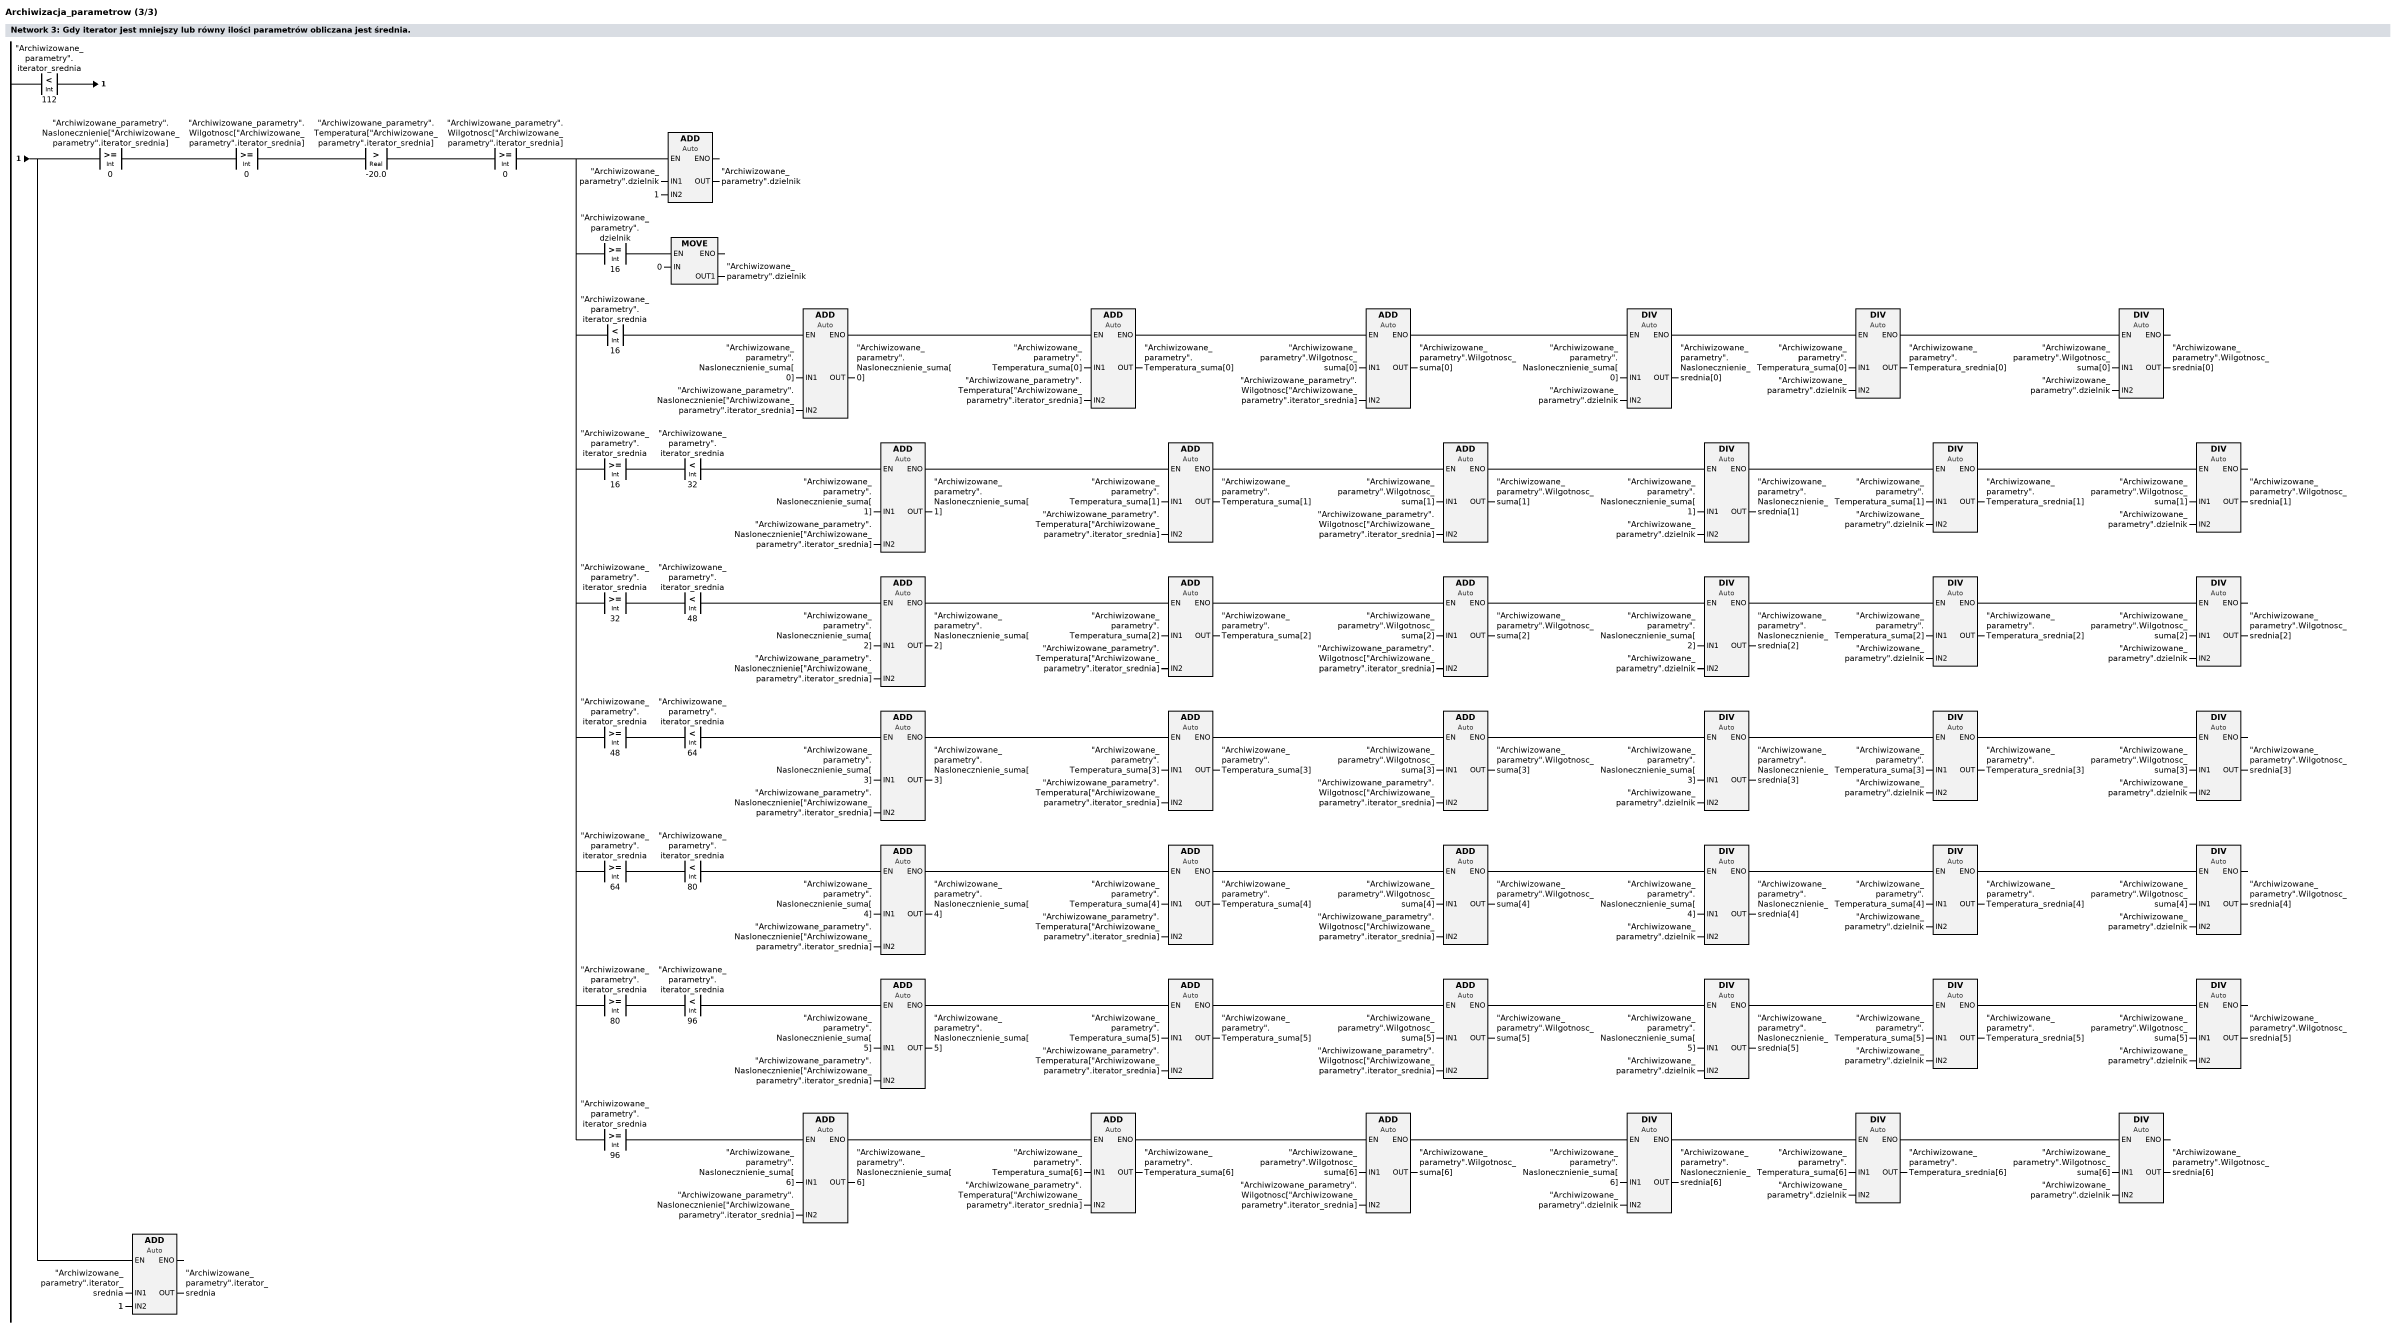
   RUNG wire#powerrail
      { S7_Templates := "SrcType := Int" } LT_Contact(in1 := "Archiwizowane_parametry".iterator_srednia, in2 := 112)
      wire#w1
      { S7_Templates := "SrcType := Int" } GE_Contact(in1 := "Archiwizowane_parametry".Naslonecznienie["Archiwizowane_parametry".iterator_srednia], in2 := 0)
      { S7_Templates := "SrcType := Int" } GE_Contact(in1 := "Archiwizowane_parametry".Wilgotnosc["Archiwizowane_parametry".iterator_srednia], in2 := 0)
      { S7_Templates := "SrcType := Real" } GT_Contact(in1 := "Archiwizowane_parametry".Temperatura["Archiwizowane_parametry".iterator_srednia], in2 := -20.0)
      { S7_Templates := "SrcType := Int" } GE_Contact(in1 := "Archiwizowane_parametry".Wilgotnosc["Archiwizowane_parametry".iterator_srednia], in2 := 0)
      wire#w2
      { S7_GenerateENO := "TRUE" } Add(in1 := "Archiwizowane_parametry".dzielnik, in2 := 1, out => "Archiwizowane_parametry".dzielnik)
   END_RUNG
   RUNG wire#w2
      { S7_Templates := "SrcType := Int" } GE_Contact(in1 := "Archiwizowane_parametry".dzielnik, in2 := 16)
      Move(in := 0, out1 => "Archiwizowane_parametry".dzielnik)
   END_RUNG
   RUNG wire#w2
      { S7_Templates := "SrcType := Int" } LT_Contact(in1 := "Archiwizowane_parametry".iterator_srednia, in2 := 16)
      { S7_GenerateENO := "TRUE" } Add(in1 := "Archiwizowane_parametry".Naslonecznienie_suma[0], in2 := "Archiwizowane_parametry".Naslonecznienie["Archiwizowane_parametry".iterator_srednia], out => "Archiwizowane_parametry".Naslonecznienie_suma[0])
      { S7_GenerateENO := "TRUE" } Add(in1 := "Archiwizowane_parametry".Temperatura_suma[0], in2 := "Archiwizowane_parametry".Temperatura["Archiwizowane_parametry".iterator_srednia], out => "Archiwizowane_parametry".Temperatura_suma[0])
      { S7_GenerateENO := "TRUE" } Add(in1 := "Archiwizowane_parametry".Wilgotnosc_suma[0], in2 := "Archiwizowane_parametry".Wilgotnosc["Archiwizowane_parametry".iterator_srednia], out => "Archiwizowane_parametry".Wilgotnosc_suma[0])
      Div(in1 := "Archiwizowane_parametry".Naslonecznienie_suma[0], in2 := "Archiwizowane_parametry".dzielnik, out => "Archiwizowane_parametry".Naslonecznienie_srednia[0])
      Div(in1 := "Archiwizowane_parametry".Temperatura_suma[0], in2 := "Archiwizowane_parametry".dzielnik, out => "Archiwizowane_parametry".Temperatura_srednia[0])
      Div(in1 := "Archiwizowane_parametry".Wilgotnosc_suma[0], in2 := "Archiwizowane_parametry".dzielnik, out => "Archiwizowane_parametry".Wilgotnosc_srednia[0])
   END_RUNG
   RUNG wire#w2
      { S7_Templates := "SrcType := Int" } GE_Contact(in1 := "Archiwizowane_parametry".iterator_srednia, in2 := 16)
      { S7_Templates := "SrcType := Int" } LT_Contact(in1 := "Archiwizowane_parametry".iterator_srednia, in2 := 32)
      { S7_GenerateENO := "TRUE" } Add(in1 := "Archiwizowane_parametry".Naslonecznienie_suma[1], in2 := "Archiwizowane_parametry".Naslonecznienie["Archiwizowane_parametry".iterator_srednia], out => "Archiwizowane_parametry".Naslonecznienie_suma[1])
      { S7_GenerateENO := "TRUE" } Add(in1 := "Archiwizowane_parametry".Temperatura_suma[1], in2 := "Archiwizowane_parametry".Temperatura["Archiwizowane_parametry".iterator_srednia], out => "Archiwizowane_parametry".Temperatura_suma[1])
      { S7_GenerateENO := "TRUE" } Add(in1 := "Archiwizowane_parametry".Wilgotnosc_suma[1], in2 := "Archiwizowane_parametry".Wilgotnosc["Archiwizowane_parametry".iterator_srednia], out => "Archiwizowane_parametry".Wilgotnosc_suma[1])
      Div(in1 := "Archiwizowane_parametry".Naslonecznienie_suma[1], in2 := "Archiwizowane_parametry".dzielnik, out => "Archiwizowane_parametry".Naslonecznienie_srednia[1])
      Div(in1 := "Archiwizowane_parametry".Temperatura_suma[1], in2 := "Archiwizowane_parametry".dzielnik, out => "Archiwizowane_parametry".Temperatura_srednia[1])
      Div(in1 := "Archiwizowane_parametry".Wilgotnosc_suma[1], in2 := "Archiwizowane_parametry".dzielnik, out => "Archiwizowane_parametry".Wilgotnosc_srednia[1])
   END_RUNG
   RUNG wire#w2
      { S7_Templates := "SrcType := Int" } GE_Contact(in1 := "Archiwizowane_parametry".iterator_srednia, in2 := 32)
      { S7_Templates := "SrcType := Int" } LT_Contact(in1 := "Archiwizowane_parametry".iterator_srednia, in2 := 48)
      { S7_GenerateENO := "TRUE" } Add(in1 := "Archiwizowane_parametry".Naslonecznienie_suma[2], in2 := "Archiwizowane_parametry".Naslonecznienie["Archiwizowane_parametry".iterator_srednia], out => "Archiwizowane_parametry".Naslonecznienie_suma[2])
      { S7_GenerateENO := "TRUE" } Add(in1 := "Archiwizowane_parametry".Temperatura_suma[2], in2 := "Archiwizowane_parametry".Temperatura["Archiwizowane_parametry".iterator_srednia], out => "Archiwizowane_parametry".Temperatura_suma[2])
      { S7_GenerateENO := "TRUE" } Add(in1 := "Archiwizowane_parametry".Wilgotnosc_suma[2], in2 := "Archiwizowane_parametry".Wilgotnosc["Archiwizowane_parametry".iterator_srednia], out => "Archiwizowane_parametry".Wilgotnosc_suma[2])
      Div(in1 := "Archiwizowane_parametry".Naslonecznienie_suma[2], in2 := "Archiwizowane_parametry".dzielnik, out => "Archiwizowane_parametry".Naslonecznienie_srednia[2])
      Div(in1 := "Archiwizowane_parametry".Temperatura_suma[2], in2 := "Archiwizowane_parametry".dzielnik, out => "Archiwizowane_parametry".Temperatura_srednia[2])
      Div(in1 := "Archiwizowane_parametry".Wilgotnosc_suma[2], in2 := "Archiwizowane_parametry".dzielnik, out => "Archiwizowane_parametry".Wilgotnosc_srednia[2])
   END_RUNG
   RUNG wire#w2
      { S7_Templates := "SrcType := Int" } GE_Contact(in1 := "Archiwizowane_parametry".iterator_srednia, in2 := 48)
      { S7_Templates := "SrcType := Int" } LT_Contact(in1 := "Archiwizowane_parametry".iterator_srednia, in2 := 64)
      { S7_GenerateENO := "TRUE" } Add(in1 := "Archiwizowane_parametry".Naslonecznienie_suma[3], in2 := "Archiwizowane_parametry".Naslonecznienie["Archiwizowane_parametry".iterator_srednia], out => "Archiwizowane_parametry".Naslonecznienie_suma[3])
      { S7_GenerateENO := "TRUE" } Add(in1 := "Archiwizowane_parametry".Temperatura_suma[3], in2 := "Archiwizowane_parametry".Temperatura["Archiwizowane_parametry".iterator_srednia], out => "Archiwizowane_parametry".Temperatura_suma[3])
      { S7_GenerateENO := "TRUE" } Add(in1 := "Archiwizowane_parametry".Wilgotnosc_suma[3], in2 := "Archiwizowane_parametry".Wilgotnosc["Archiwizowane_parametry".iterator_srednia], out => "Archiwizowane_parametry".Wilgotnosc_suma[3])
      Div(in1 := "Archiwizowane_parametry".Naslonecznienie_suma[3], in2 := "Archiwizowane_parametry".dzielnik, out => "Archiwizowane_parametry".Naslonecznienie_srednia[3])
      Div(in1 := "Archiwizowane_parametry".Temperatura_suma[3], in2 := "Archiwizowane_parametry".dzielnik, out => "Archiwizowane_parametry".Temperatura_srednia[3])
      Div(in1 := "Archiwizowane_parametry".Wilgotnosc_suma[3], in2 := "Archiwizowane_parametry".dzielnik, out => "Archiwizowane_parametry".Wilgotnosc_srednia[3])
   END_RUNG
   RUNG wire#w2
      { S7_Templates := "SrcType := Int" } GE_Contact(in1 := "Archiwizowane_parametry".iterator_srednia, in2 := 64)
      { S7_Templates := "SrcType := Int" } LT_Contact(in1 := "Archiwizowane_parametry".iterator_srednia, in2 := 80)
      { S7_GenerateENO := "TRUE" } Add(in1 := "Archiwizowane_parametry".Naslonecznienie_suma[4], in2 := "Archiwizowane_parametry".Naslonecznienie["Archiwizowane_parametry".iterator_srednia], out => "Archiwizowane_parametry".Naslonecznienie_suma[4])
      { S7_GenerateENO := "TRUE" } Add(in1 := "Archiwizowane_parametry".Temperatura_suma[4], in2 := "Archiwizowane_parametry".Temperatura["Archiwizowane_parametry".iterator_srednia], out => "Archiwizowane_parametry".Temperatura_suma[4])
      { S7_GenerateENO := "TRUE" } Add(in1 := "Archiwizowane_parametry".Wilgotnosc_suma[4], in2 := "Archiwizowane_parametry".Wilgotnosc["Archiwizowane_parametry".iterator_srednia], out => "Archiwizowane_parametry".Wilgotnosc_suma[4])
      Div(in1 := "Archiwizowane_parametry".Naslonecznienie_suma[4], in2 := "Archiwizowane_parametry".dzielnik, out => "Archiwizowane_parametry".Naslonecznienie_srednia[4])
      Div(in1 := "Archiwizowane_parametry".Temperatura_suma[4], in2 := "Archiwizowane_parametry".dzielnik, out => "Archiwizowane_parametry".Temperatura_srednia[4])
      Div(in1 := "Archiwizowane_parametry".Wilgotnosc_suma[4], in2 := "Archiwizowane_parametry".dzielnik, out => "Archiwizowane_parametry".Wilgotnosc_srednia[4])
   END_RUNG
   RUNG wire#w2
      { S7_Templates := "SrcType := Int" } GE_Contact(in1 := "Archiwizowane_parametry".iterator_srednia, in2 := 80)
      { S7_Templates := "SrcType := Int" } LT_Contact(in1 := "Archiwizowane_parametry".iterator_srednia, in2 := 96)
      { S7_GenerateENO := "TRUE" } Add(in1 := "Archiwizowane_parametry".Naslonecznienie_suma[5], in2 := "Archiwizowane_parametry".Naslonecznienie["Archiwizowane_parametry".iterator_srednia], out => "Archiwizowane_parametry".Naslonecznienie_suma[5])
      { S7_GenerateENO := "TRUE" } Add(in1 := "Archiwizowane_parametry".Temperatura_suma[5], in2 := "Archiwizowane_parametry".Temperatura["Archiwizowane_parametry".iterator_srednia], out => "Archiwizowane_parametry".Temperatura_suma[5])
      { S7_GenerateENO := "TRUE" } Add(in1 := "Archiwizowane_parametry".Wilgotnosc_suma[5], in2 := "Archiwizowane_parametry".Wilgotnosc["Archiwizowane_parametry".iterator_srednia], out => "Archiwizowane_parametry".Wilgotnosc_suma[5])
      Div(in1 := "Archiwizowane_parametry".Naslonecznienie_suma[5], in2 := "Archiwizowane_parametry".dzielnik, out => "Archiwizowane_parametry".Naslonecznienie_srednia[5])
      Div(in1 := "Archiwizowane_parametry".Temperatura_suma[5], in2 := "Archiwizowane_parametry".dzielnik, out => "Archiwizowane_parametry".Temperatura_srednia[5])
      Div(in1 := "Archiwizowane_parametry".Wilgotnosc_suma[5], in2 := "Archiwizowane_parametry".dzielnik, out => "Archiwizowane_parametry".Wilgotnosc_srednia[5])
   END_RUNG
   RUNG wire#w2
      { S7_Templates := "SrcType := Int" } GE_Contact(in1 := "Archiwizowane_parametry".iterator_srednia, in2 := 96)
      { S7_GenerateENO := "TRUE" } Add(in1 := "Archiwizowane_parametry".Naslonecznienie_suma[6], in2 := "Archiwizowane_parametry".Naslonecznienie["Archiwizowane_parametry".iterator_srednia], out => "Archiwizowane_parametry".Naslonecznienie_suma[6])
      { S7_GenerateENO := "TRUE" } Add(in1 := "Archiwizowane_parametry".Temperatura_suma[6], in2 := "Archiwizowane_parametry".Temperatura["Archiwizowane_parametry".iterator_srednia], out => "Archiwizowane_parametry".Temperatura_suma[6])
      { S7_GenerateENO := "TRUE" } Add(in1 := "Archiwizowane_parametry".Wilgotnosc_suma[6], in2 := "Archiwizowane_parametry".Wilgotnosc["Archiwizowane_parametry".iterator_srednia], out => "Archiwizowane_parametry".Wilgotnosc_suma[6])
      Div(in1 := "Archiwizowane_parametry".Naslonecznienie_suma[6], in2 := "Archiwizowane_parametry".dzielnik, out => "Archiwizowane_parametry".Naslonecznienie_srednia[6])
      Div(in1 := "Archiwizowane_parametry".Temperatura_suma[6], in2 := "Archiwizowane_parametry".dzielnik, out => "Archiwizowane_parametry".Temperatura_srednia[6])
      Div(in1 := "Archiwizowane_parametry".Wilgotnosc_suma[6], in2 := "Archiwizowane_parametry".dzielnik, out => "Archiwizowane_parametry".Wilgotnosc_srednia[6])
   END_RUNG
   RUNG wire#w1
      { S7_GenerateENO := "TRUE" } Add(in1 := "Archiwizowane_parametry".iterator_srednia, in2 := 1, out => "Archiwizowane_parametry".iterator_srednia)
   END_RUNG
   // the same network as SCL:
   // ENO of a box is taken as its EN; it also drops when the box reports an error
   #_w1 := "Archiwizowane_parametry".iterator_srednia < 112;
   #_w2 := #_w1 AND ("Archiwizowane_parametry".Naslonecznienie["Archiwizowane_parametry".iterator_srednia] >= 0) AND ("Archiwizowane_parametry".Wilgotnosc["Archiwizowane_parametry".iterator_srednia] >= 0) AND ("Archiwizowane_parametry".Temperatura["Archiwizowane_parametry".iterator_srednia] > (-20.0)) AND ("Archiwizowane_parametry".Wilgotnosc["Archiwizowane_parametry".iterator_srednia] >= 0);
   IF #_w2 THEN "Archiwizowane_parametry".dzielnik := "Archiwizowane_parametry".dzielnik + 1; END_IF;
   IF #_w2 AND ("Archiwizowane_parametry".dzielnik >= 16) THEN
       "Archiwizowane_parametry".dzielnik := 0;
   END_IF;
   IF #_w2 AND ("Archiwizowane_parametry".iterator_srednia < 16) THEN
       "Archiwizowane_parametry".Naslonecznienie_suma[0] := "Archiwizowane_parametry".Naslonecznienie_suma[0] + "Archiwizowane_parametry".Naslonecznienie["Archiwizowane_parametry".iterator_srednia];
       "Archiwizowane_parametry".Temperatura_suma[0] := "Archiwizowane_parametry".Temperatura_suma[0] + "Archiwizowane_parametry".Temperatura["Archiwizowane_parametry".iterator_srednia];
       "Archiwizowane_parametry".Wilgotnosc_suma[0] := "Archiwizowane_parametry".Wilgotnosc_suma[0] + "Archiwizowane_parametry".Wilgotnosc["Archiwizowane_parametry".iterator_srednia];
       "Archiwizowane_parametry".Naslonecznienie_srednia[0] := "Archiwizowane_parametry".Naslonecznienie_suma[0] / "Archiwizowane_parametry".dzielnik;
       "Archiwizowane_parametry".Temperatura_srednia[0] := "Archiwizowane_parametry".Temperatura_suma[0] / "Archiwizowane_parametry".dzielnik;
       "Archiwizowane_parametry".Wilgotnosc_srednia[0] := "Archiwizowane_parametry".Wilgotnosc_suma[0] / "Archiwizowane_parametry".dzielnik;
   END_IF;
   IF #_w2 AND ("Archiwizowane_parametry".iterator_srednia >= 16) AND ("Archiwizowane_parametry".iterator_srednia < 32) THEN
       "Archiwizowane_parametry".Naslonecznienie_suma[1] := "Archiwizowane_parametry".Naslonecznienie_suma[1] + "Archiwizowane_parametry".Naslonecznienie["Archiwizowane_parametry".iterator_srednia];
       "Archiwizowane_parametry".Temperatura_suma[1] := "Archiwizowane_parametry".Temperatura_suma[1] + "Archiwizowane_parametry".Temperatura["Archiwizowane_parametry".iterator_srednia];
       "Archiwizowane_parametry".Wilgotnosc_suma[1] := "Archiwizowane_parametry".Wilgotnosc_suma[1] + "Archiwizowane_parametry".Wilgotnosc["Archiwizowane_parametry".iterator_srednia];
       "Archiwizowane_parametry".Naslonecznienie_srednia[1] := "Archiwizowane_parametry".Naslonecznienie_suma[1] / "Archiwizowane_parametry".dzielnik;
       "Archiwizowane_parametry".Temperatura_srednia[1] := "Archiwizowane_parametry".Temperatura_suma[1] / "Archiwizowane_parametry".dzielnik;
       "Archiwizowane_parametry".Wilgotnosc_srednia[1] := "Archiwizowane_parametry".Wilgotnosc_suma[1] / "Archiwizowane_parametry".dzielnik;
   END_IF;
   IF #_w2 AND ("Archiwizowane_parametry".iterator_srednia >= 32) AND ("Archiwizowane_parametry".iterator_srednia < 48) THEN
       "Archiwizowane_parametry".Naslonecznienie_suma[2] := "Archiwizowane_parametry".Naslonecznienie_suma[2] + "Archiwizowane_parametry".Naslonecznienie["Archiwizowane_parametry".iterator_srednia];
       "Archiwizowane_parametry".Temperatura_suma[2] := "Archiwizowane_parametry".Temperatura_suma[2] + "Archiwizowane_parametry".Temperatura["Archiwizowane_parametry".iterator_srednia];
       "Archiwizowane_parametry".Wilgotnosc_suma[2] := "Archiwizowane_parametry".Wilgotnosc_suma[2] + "Archiwizowane_parametry".Wilgotnosc["Archiwizowane_parametry".iterator_srednia];
       "Archiwizowane_parametry".Naslonecznienie_srednia[2] := "Archiwizowane_parametry".Naslonecznienie_suma[2] / "Archiwizowane_parametry".dzielnik;
       "Archiwizowane_parametry".Temperatura_srednia[2] := "Archiwizowane_parametry".Temperatura_suma[2] / "Archiwizowane_parametry".dzielnik;
       "Archiwizowane_parametry".Wilgotnosc_srednia[2] := "Archiwizowane_parametry".Wilgotnosc_suma[2] / "Archiwizowane_parametry".dzielnik;
   END_IF;
   IF #_w2 AND ("Archiwizowane_parametry".iterator_srednia >= 48) AND ("Archiwizowane_parametry".iterator_srednia < 64) THEN
       "Archiwizowane_parametry".Naslonecznienie_suma[3] := "Archiwizowane_parametry".Naslonecznienie_suma[3] + "Archiwizowane_parametry".Naslonecznienie["Archiwizowane_parametry".iterator_srednia];
       "Archiwizowane_parametry".Temperatura_suma[3] := "Archiwizowane_parametry".Temperatura_suma[3] + "Archiwizowane_parametry".Temperatura["Archiwizowane_parametry".iterator_srednia];
       "Archiwizowane_parametry".Wilgotnosc_suma[3] := "Archiwizowane_parametry".Wilgotnosc_suma[3] + "Archiwizowane_parametry".Wilgotnosc["Archiwizowane_parametry".iterator_srednia];
       "Archiwizowane_parametry".Naslonecznienie_srednia[3] := "Archiwizowane_parametry".Naslonecznienie_suma[3] / "Archiwizowane_parametry".dzielnik;
       "Archiwizowane_parametry".Temperatura_srednia[3] := "Archiwizowane_parametry".Temperatura_suma[3] / "Archiwizowane_parametry".dzielnik;
       "Archiwizowane_parametry".Wilgotnosc_srednia[3] := "Archiwizowane_parametry".Wilgotnosc_suma[3] / "Archiwizowane_parametry".dzielnik;
   END_IF;
   IF #_w2 AND ("Archiwizowane_parametry".iterator_srednia >= 64) AND ("Archiwizowane_parametry".iterator_srednia < 80) THEN
       "Archiwizowane_parametry".Naslonecznienie_suma[4] := "Archiwizowane_parametry".Naslonecznienie_suma[4] + "Archiwizowane_parametry".Naslonecznienie["Archiwizowane_parametry".iterator_srednia];
       "Archiwizowane_parametry".Temperatura_suma[4] := "Archiwizowane_parametry".Temperatura_suma[4] + "Archiwizowane_parametry".Temperatura["Archiwizowane_parametry".iterator_srednia];
       "Archiwizowane_parametry".Wilgotnosc_suma[4] := "Archiwizowane_parametry".Wilgotnosc_suma[4] + "Archiwizowane_parametry".Wilgotnosc["Archiwizowane_parametry".iterator_srednia];
       "Archiwizowane_parametry".Naslonecznienie_srednia[4] := "Archiwizowane_parametry".Naslonecznienie_suma[4] / "Archiwizowane_parametry".dzielnik;
       "Archiwizowane_parametry".Temperatura_srednia[4] := "Archiwizowane_parametry".Temperatura_suma[4] / "Archiwizowane_parametry".dzielnik;
       "Archiwizowane_parametry".Wilgotnosc_srednia[4] := "Archiwizowane_parametry".Wilgotnosc_suma[4] / "Archiwizowane_parametry".dzielnik;
   END_IF;
   IF #_w2 AND ("Archiwizowane_parametry".iterator_srednia >= 80) AND ("Archiwizowane_parametry".iterator_srednia < 96) THEN
       "Archiwizowane_parametry".Naslonecznienie_suma[5] := "Archiwizowane_parametry".Naslonecznienie_suma[5] + "Archiwizowane_parametry".Naslonecznienie["Archiwizowane_parametry".iterator_srednia];
       "Archiwizowane_parametry".Temperatura_suma[5] := "Archiwizowane_parametry".Temperatura_suma[5] + "Archiwizowane_parametry".Temperatura["Archiwizowane_parametry".iterator_srednia];
       "Archiwizowane_parametry".Wilgotnosc_suma[5] := "Archiwizowane_parametry".Wilgotnosc_suma[5] + "Archiwizowane_parametry".Wilgotnosc["Archiwizowane_parametry".iterator_srednia];
       "Archiwizowane_parametry".Naslonecznienie_srednia[5] := "Archiwizowane_parametry".Naslonecznienie_suma[5] / "Archiwizowane_parametry".dzielnik;
       "Archiwizowane_parametry".Temperatura_srednia[5] := "Archiwizowane_parametry".Temperatura_suma[5] / "Archiwizowane_parametry".dzielnik;
       "Archiwizowane_parametry".Wilgotnosc_srednia[5] := "Archiwizowane_parametry".Wilgotnosc_suma[5] / "Archiwizowane_parametry".dzielnik;
   END_IF;
   IF #_w2 AND ("Archiwizowane_parametry".iterator_srednia >= 96) THEN
       "Archiwizowane_parametry".Naslonecznienie_suma[6] := "Archiwizowane_parametry".Naslonecznienie_suma[6] + "Archiwizowane_parametry".Naslonecznienie["Archiwizowane_parametry".iterator_srednia];
       "Archiwizowane_parametry".Temperatura_suma[6] := "Archiwizowane_parametry".Temperatura_suma[6] + "Archiwizowane_parametry".Temperatura["Archiwizowane_parametry".iterator_srednia];
       "Archiwizowane_parametry".Wilgotnosc_suma[6] := "Archiwizowane_parametry".Wilgotnosc_suma[6] + "Archiwizowane_parametry".Wilgotnosc["Archiwizowane_parametry".iterator_srednia];
       "Archiwizowane_parametry".Naslonecznienie_srednia[6] := "Archiwizowane_parametry".Naslonecznienie_suma[6] / "Archiwizowane_parametry".dzielnik;
       "Archiwizowane_parametry".Temperatura_srednia[6] := "Archiwizowane_parametry".Temperatura_suma[6] / "Archiwizowane_parametry".dzielnik;
       "Archiwizowane_parametry".Wilgotnosc_srednia[6] := "Archiwizowane_parametry".Wilgotnosc_suma[6] / "Archiwizowane_parametry".dzielnik;
   END_IF;
   IF #_w1 THEN
       "Archiwizowane_parametry".iterator_srednia := "Archiwizowane_parametry".iterator_srednia + 1;
   END_IF;
END_REGION
END_FUNCTION

// folder: LGF/4 Math operations

FUNCTION "LGF_RandomRange_Real" : Real   // FC10014, SCL
TITLE = LGF_RandomRange_Real
{ S7_Optimized_Access := 'TRUE' }
AUTHOR : Siemens_Digital_Industries
FAMILY : LGF
NAME : LGF_RandomRange_Real
// This function generates random numbers in defined limits (Datatype Real)
   VAR_INPUT
      minValue : Real;   // minimal Value random can reach / Minimum value of the range of the random number
      maxValue : Real;   // maximal Value random can reach / Maximum value of the range of the random number
   END_VAR
   VAR_OUTPUT
      error : Bool;   // Error if true
      status : Word;   // Status of the function
      subfunctionStatus : Word;   // Status or return value of called FB's, FCs and system blocks
   END_VAR
   VAR_TEMP
      tempTime : DTL;   // System time
      tempNanoSecondInDWord : DWord;   // UDINT converted to DWORD for access to individual bytes
      tempTimeStatus : Word;   // Status of the instruction RD_SYS_T
      tempRandomValue : DWord;   // Random-start-value
      tempNormReal : Real;   // normalized value
   END_VAR
   // Ret_Val : Returns random Real number in predefined range
   VAR CONSTANT
      ZERO : Real := 0.0;   // Zero value in case of error
      MAX_UDINT : UDInt := 4294967295;   // Maximum UDINT value
      SUB_STATUS_NO_ERROR : Word := 16#0000;   // Status: sub function call ends without error
      STATUS_FINISHED_NO_ERROR : Word := 16#0000;   // Status: Execution finished without errors
      ERR_MAX_LESS_MIN : Word := 16#8200;   // Error: The maximum limit number is smaller than the minimum limit number
      ERR_RD_SYS_T : Word := 16#8600;   // Error: System function Read system time returned an error
   END_VAR
BEGIN
   REGION Block info header
     //=============================================================================
     // SIEMENS AG / (c)Copyright 2017
     //-----------------------------------------------------------------------------
     // Title:            LGF_RandomRange_Real
     // Comment/Function: This function generates random numbers in defined limits (Datatype Real)
     // Library/Family:   LGF(Library General Functions)
     // Author:           Siemens Digital Industry Support
     // Tested with:      S7-PLCSIM Advanced V2.0 SP1
     // Engineering:      TIA Portal V15 Update 2
     // Restrictions:     ENO disabled - error handling done by error and status
     // Requirements:     PLC (S7-1200 / S7-1500)
     //-------------------------------------------------------------------------------
     // Change log table:
     // Version  | Date       | Expert in charge       | Changes applied
     //----------|------------|------------------------|------------------------------
     // 01.00.00 19.08.2015  Siemens Industry Online Support
     //                      First released version
     // 01.00.01 02.01.2017  Siemens Industry Online Support
     //                      Upgrade: TIA Portal V14 Update 1
     // 01.00.02 02.03.2017  Siemens Industry Online Support
     //                      Bugfix: FC number
     // 01.00.03 17.08.2018  Siemens Industry Online Support
     //                      Upgrade: TIA V15 Update 2
     // 01.00.04 23.11.2018  Siemens Industry Online Support
     //                      Upgrade: TIA V15.1
     // 01.01.00 13.11.2019  Siemens Industry Presales Support
     //                      Renamed from "LGF_RandomReal" to "LGF_RandomRange_Real"
     //                      Regions, commens and costants are added
     // 03.00.00 23.04.2020  Siemens Industry Support
     //                      Set version to V3.0.0, harmonize the version of the whole library
     //=============================================================================
   END_REGION

   REGION Validation
     // Check if the maximal Value is less than the minimal value
     IF (#minValue > #maxValue) THEN
       #error := true;
       #status := #ERR_MAX_LESS_MIN;
       #subfunctionStatus := #SUB_STATUS_NO_ERROR;
       #LGF_RandomRange_Real := #ZERO;
       RETURN;
     END_IF;

     // Read system time
     #tempTimeStatus := INT_TO_WORD(RD_SYS_T(#tempTime));

     // Check return variable for error
     IF (#tempTimeStatus <> #SUB_STATUS_NO_ERROR) THEN
       #error := true;
       #status := #ERR_RD_SYS_T;
       #subfunctionStatus := #tempTimeStatus;
       #LGF_RandomRange_Real := #ZERO;
       RETURN;
     END_IF;
   END_REGION

   REGION Calculating random number
     // Converting to double word so individual bytes can be addressed
     #tempNanoSecondInDWord := UDINT_TO_DWORD(#tempTime.NANOSECOND);

     // Calculate a random-start-value depending on the time
     #tempRandomValue.%B3 := #tempNanoSecondInDWord.%B0;
     #tempRandomValue.%B2 := #tempNanoSecondInDWord.%B1;
     #tempRandomValue.%B1 := #tempNanoSecondInDWord.%B2;
     #tempRandomValue.%B0 := #tempNanoSecondInDWord.%B3;

     // Norm the calculated random number: 0.0 <= #tempNormReal <= 1.0
     #tempNormReal := UDINT_TO_REAL(DWORD_TO_UDINT(#tempRandomValue)) / UDINT_TO_REAL(#MAX_UDINT);

     // Scale the tempNormReal to be in the range of maxValue and minValue
     #LGF_RandomRange_Real := ((#tempNormReal * (#maxValue - #minValue) + (#minValue)));

     #error := false;
     #status := #STATUS_FINISHED_NO_ERROR;
     #subfunctionStatus := #SUB_STATUS_NO_ERROR;
     // ENO mechanism is not used
     ENO := TRUE;
   END_REGION
END_FUNCTION

// ===== PLC "PLC_Web_server"  CPU 1518-4 PN/DP =====

VAR_GLOBAL   // PLC tag table "Default tag table"
   "err" AT %MW1 : Int;
   "tag1" AT %M6.0 : Bool;
END_VAR

DATA_BLOCK "Wejscia_PLC"   // DB2
{ S7_Optimized_Access := 'TRUE' }
VERSION : 0.1
   VAR
      Czujnik_wilgotności_powietrza : Int;   // Czujnik wilgotności powietrza w szklarni
      Czujnik_wilgotności_gleby : Int;   // Czujnik wilgotności gleby w szklarni
      Temperatura_wewnetrzna : Real;   // Temperatura wewnątrz szklarni
      Czujnik_natezenia_swiatła : Int;   // Czujnik natężenia światła wewnątrz szklarni
      Wewnetrzny_czujnik_CO2 : Int;   // Czujnik stężenia dwutlenku węgla w szklarni
      Stopien_zasloniecia_rolet : Int;   // Stopień zasłonięcia rolet w szklarni (przyjęty przedział 0-100%)
   END_VAR
BEGIN
END_DATA_BLOCK

// folder: Archiwizacja_parametrow

DATA_BLOCK "Archiwizowane_parametry"   // DB4
{ S7_Optimized_Access := 'TRUE' }
VERSION : 0.1
   VAR
      Temperatura : Array[0..111] of Real;
      Wilgotnosc : Array[0..111] of Int;
      Naslonecznienie : Array[0..111] of Int;
      iterator : Int := 0;   // Iterator służący do zapisu danych w odpowiednich komórkach tablicy.
      Temperatura_srednia : Array[0..6] of Real;
      Wilgotnosc_srednia : Array[0..6] of Int;
      Naslonecznienie_srednia : Array[0..6] of Int;
      iterator_srednia : Int := 0;   // Iterator służący do zapisu danych w odpowiednich komórkach tablicy.
      dzielnik : Int;   // Ilość zsumowanych parametrów w średniej
      Temperatura_suma : Array[0..6] of Real;
      Wilgotnosc_suma : Array[0..6] of Int;
      Naslonecznienie_suma : Array[0..6] of Int;
   END_VAR
BEGIN
   Naslonecznienie[0] := -1;
   Naslonecznienie[1] := -1;
   Temperatura[0] := -20.0;
   Temperatura[1] := -20.0;
   Temperatura[2] := -20.0;
   Temperatura[3] := -20.0;
   Temperatura[4] := -20.0;
   Temperatura[5] := -20.0;
   Temperatura[12] := -20.0;
   Temperatura[13] := -20.0;
   Temperatura[14] := -20.0;
   Temperatura[15] := -20.0;
   Temperatura[16] := -20.0;
   Temperatura[17] := -20.0;
   Temperatura[6] := -20.0;
   Temperatura[7] := -20.0;
   Temperatura[8] := -20.0;
   Temperatura[9] := -20.0;
   Temperatura[10] := -20.0;
   Temperatura[11] := -20.0;
   Temperatura[18] := -20.0;
   Temperatura[19] := -20.0;
   Temperatura[20] := -20.0;
   Temperatura[21] := -20.0;
   Temperatura[22] := -20.0;
   Temperatura[23] := -20.0;
   Temperatura[24] := -20.0;
   Temperatura[25] := -20.0;
   Temperatura[26] := -20.0;
   Temperatura[27] := -20.0;
   Temperatura[28] := -20.0;
   Temperatura[29] := -20.0;
   Temperatura[30] := -20.0;
   Temperatura[31] := -20.0;
   Temperatura[32] := -20.0;
   Temperatura[33] := -20.0;
   Temperatura[34] := -20.0;
   Temperatura[35] := -20.0;
   Temperatura[36] := -20.0;
   Temperatura[37] := -20.0;
   Temperatura[38] := -20.0;
   Temperatura[39] := -20.0;
   Temperatura[40] := -20.0;
   Temperatura[41] := -20.0;
   Temperatura[42] := -20.0;
   Temperatura[43] := -20.0;
   Temperatura[44] := -20.0;
   Temperatura[45] := -20.0;
   Temperatura[46] := -20.0;
   Temperatura[47] := -20.0;
   Temperatura[48] := -20.0;
   Temperatura[49] := -20.0;
   Temperatura[50] := -20.0;
   Temperatura[51] := -20.0;
   Temperatura[52] := -20.0;
   Temperatura[53] := -20.0;
   Temperatura[54] := -20.0;
   Temperatura[55] := -20.0;
   Temperatura[56] := -20.0;
   Temperatura[57] := -20.0;
   Temperatura[58] := -20.0;
   Temperatura[59] := -20.0;
   Temperatura[60] := -20.0;
   Temperatura[61] := -20.0;
   Temperatura[62] := -20.0;
   Temperatura[63] := -20.0;
   Temperatura[64] := -20.0;
   Temperatura[65] := -20.0;
   Temperatura[66] := -20.0;
   Temperatura[67] := -20.0;
   Temperatura[68] := -20.0;
   Temperatura[69] := -20.0;
   Temperatura[70] := -20.0;
   Temperatura[71] := -20.0;
   Temperatura[72] := -20.0;
   Temperatura[73] := -20.0;
   Temperatura[74] := -20.0;
   Temperatura[75] := -20.0;
   Temperatura[76] := -20.0;
   Temperatura[77] := -20.0;
   Temperatura[78] := -20.0;
   Temperatura[79] := -20.0;
   Temperatura[80] := -20.0;
   Temperatura[81] := -20.0;
   Temperatura[82] := -20.0;
   Temperatura[83] := -20.0;
   Temperatura[84] := -20.0;
   Temperatura[85] := -20.0;
   Temperatura[86] := -20.0;
   Temperatura[87] := -20.0;
   Temperatura[88] := -20.0;
   Temperatura[89] := -20.0;
   Temperatura[90] := -20.0;
   Temperatura[91] := -20.0;
   Temperatura[92] := -20.0;
   Temperatura[93] := -20.0;
   Temperatura[94] := -20.0;
   Temperatura[95] := -20.0;
   Temperatura[96] := -20.0;
   Temperatura[97] := -20.0;
   Temperatura[98] := -20.0;
   Temperatura[99] := -20.0;
   Temperatura[100] := -20.0;
   Temperatura[101] := -20.0;
   Temperatura[102] := -20.0;
   Temperatura[103] := -20.0;
   Temperatura[104] := -20.0;
   Temperatura[105] := -20.0;
   Temperatura[106] := -20.0;
   Temperatura[107] := -20.0;
   Temperatura[108] := -20.0;
   Temperatura[109] := -20.0;
   Temperatura[110] := -20.0;
   Temperatura[111] := -20.0;
   Wilgotnosc[0] := -1;
   Wilgotnosc[1] := -1;
   Wilgotnosc[2] := -1;
   Wilgotnosc[3] := -1;
   Wilgotnosc[4] := -1;
   Wilgotnosc[5] := -1;
   Wilgotnosc[6] := -1;
   Wilgotnosc[7] := -1;
   Wilgotnosc[8] := -1;
   Wilgotnosc[9] := -1;
   Wilgotnosc[10] := -1;
   Wilgotnosc[11] := -1;
   Wilgotnosc[12] := -1;
   Wilgotnosc[13] := -1;
   Wilgotnosc[14] := -1;
   Wilgotnosc[15] := -1;
   Wilgotnosc[16] := -1;
   Wilgotnosc[17] := -1;
   Wilgotnosc[18] := -1;
   Wilgotnosc[19] := -1;
   Wilgotnosc[20] := -1;
   Wilgotnosc[21] := -1;
   Wilgotnosc[22] := -1;
   Wilgotnosc[23] := -1;
   Wilgotnosc[24] := -1;
   Wilgotnosc[25] := -1;
   Wilgotnosc[26] := -1;
   Wilgotnosc[27] := -1;
   Wilgotnosc[28] := -1;
   Wilgotnosc[29] := -1;
   Wilgotnosc[30] := -1;
   Wilgotnosc[31] := -1;
   Wilgotnosc[32] := -1;
   Wilgotnosc[33] := -1;
   Wilgotnosc[34] := -1;
   Wilgotnosc[35] := -1;
   Wilgotnosc[36] := -1;
   Wilgotnosc[37] := -1;
   Wilgotnosc[38] := -1;
   Wilgotnosc[39] := -1;
   Wilgotnosc[40] := -1;
   Wilgotnosc[41] := -1;
   Wilgotnosc[42] := -1;
   Wilgotnosc[43] := -1;
   Wilgotnosc[44] := -1;
   Wilgotnosc[45] := -1;
   Wilgotnosc[46] := -1;
   Wilgotnosc[47] := -1;
   Wilgotnosc[48] := -1;
   Wilgotnosc[49] := -1;
   Wilgotnosc[50] := -1;
   Wilgotnosc[51] := -1;
   Wilgotnosc[52] := -1;
   Wilgotnosc[53] := -1;
   Wilgotnosc[54] := -1;
   Wilgotnosc[55] := -1;
   Wilgotnosc[56] := -1;
   Wilgotnosc[57] := -1;
   Wilgotnosc[58] := -1;
   Wilgotnosc[59] := -1;
   Wilgotnosc[60] := -1;
   Wilgotnosc[61] := -1;
   Wilgotnosc[62] := -1;
   Wilgotnosc[63] := -1;
   Wilgotnosc[64] := -1;
   Wilgotnosc[65] := -1;
   Wilgotnosc[66] := -1;
   Wilgotnosc[67] := -1;
   Wilgotnosc[68] := -1;
   Wilgotnosc[69] := -1;
   Wilgotnosc[70] := -1;
   Wilgotnosc[71] := -1;
   Wilgotnosc[72] := -1;
   Wilgotnosc[73] := -1;
   Wilgotnosc[74] := -1;
   Wilgotnosc[75] := -1;
   Wilgotnosc[76] := -1;
   Wilgotnosc[77] := -1;
   Wilgotnosc[78] := -1;
   Wilgotnosc[79] := -1;
   Wilgotnosc[80] := -1;
   Wilgotnosc[81] := -1;
   Wilgotnosc[82] := -1;
   Wilgotnosc[83] := -1;
   Wilgotnosc[84] := -1;
   Wilgotnosc[85] := -1;
   Wilgotnosc[86] := -1;
   Wilgotnosc[87] := -1;
   Wilgotnosc[88] := -1;
   Wilgotnosc[89] := -1;
   Wilgotnosc[90] := -1;
   Wilgotnosc[91] := -1;
   Wilgotnosc[92] := -1;
   Wilgotnosc[93] := -1;
   Wilgotnosc[94] := -1;
   Wilgotnosc[95] := -1;
   Wilgotnosc[96] := -1;
   Wilgotnosc[97] := -1;
   Wilgotnosc[98] := -1;
   Wilgotnosc[99] := -1;
   Wilgotnosc[100] := -1;
   Wilgotnosc[101] := -1;
   Wilgotnosc[102] := -1;
   Wilgotnosc[103] := -1;
   Wilgotnosc[104] := -1;
   Wilgotnosc[105] := -1;
   Wilgotnosc[106] := -1;
   Wilgotnosc[107] := -1;
   Wilgotnosc[108] := -1;
   Wilgotnosc[109] := -1;
   Wilgotnosc[110] := -1;
   Wilgotnosc[111] := -1;
   Naslonecznienie[2] := -1;
   Naslonecznienie[3] := -1;
   Naslonecznienie[4] := -1;
   Naslonecznienie[5] := -1;
   Naslonecznienie[6] := -1;
   Naslonecznienie[7] := -1;
   Naslonecznienie[8] := -1;
   Naslonecznienie[9] := -1;
   Naslonecznienie[10] := -1;
   Naslonecznienie[11] := -1;
   Naslonecznienie[12] := -1;
   Naslonecznienie[13] := -1;
   Naslonecznienie[14] := -1;
   Naslonecznienie[15] := -1;
   Naslonecznienie[16] := -1;
   Naslonecznienie[17] := -1;
   Naslonecznienie[18] := -1;
   Naslonecznienie[19] := -1;
   Naslonecznienie[20] := -1;
   Naslonecznienie[21] := -1;
   Naslonecznienie[22] := -1;
   Naslonecznienie[23] := -1;
   Naslonecznienie[24] := -1;
   Naslonecznienie[25] := -1;
   Naslonecznienie[26] := -1;
   Naslonecznienie[27] := -1;
   Naslonecznienie[28] := -1;
   Naslonecznienie[29] := -1;
   Naslonecznienie[30] := -1;
   Naslonecznienie[31] := -1;
   Naslonecznienie[32] := -1;
   Naslonecznienie[33] := -1;
   Naslonecznienie[34] := -1;
   Naslonecznienie[35] := -1;
   Naslonecznienie[36] := -1;
   Naslonecznienie[37] := -1;
   Naslonecznienie[38] := -1;
   Naslonecznienie[39] := -1;
   Naslonecznienie[40] := -1;
   Naslonecznienie[41] := -1;
   Naslonecznienie[42] := -1;
   Naslonecznienie[43] := -1;
   Naslonecznienie[44] := -1;
   Naslonecznienie[45] := -1;
   Naslonecznienie[46] := -1;
   Naslonecznienie[47] := -1;
   Naslonecznienie[48] := -1;
   Naslonecznienie[49] := -1;
   Naslonecznienie[50] := -1;
   Naslonecznienie[51] := -1;
   Naslonecznienie[52] := -1;
   Naslonecznienie[53] := -1;
   Naslonecznienie[54] := -1;
   Naslonecznienie[55] := -1;
   Naslonecznienie[56] := -1;
   Naslonecznienie[57] := -1;
   Naslonecznienie[58] := -1;
   Naslonecznienie[59] := -1;
   Naslonecznienie[60] := -1;
   Naslonecznienie[61] := -1;
   Naslonecznienie[62] := -1;
   Naslonecznienie[63] := -1;
   Naslonecznienie[64] := -1;
   Naslonecznienie[65] := -1;
   Naslonecznienie[66] := -1;
   Naslonecznienie[67] := -1;
   Naslonecznienie[68] := -1;
   Naslonecznienie[69] := -1;
   Naslonecznienie[70] := -1;
   Naslonecznienie[71] := -1;
   Naslonecznienie[72] := -1;
   Naslonecznienie[73] := -1;
   Naslonecznienie[74] := -1;
   Naslonecznienie[75] := -1;
   Naslonecznienie[76] := -1;
   Naslonecznienie[77] := -1;
   Naslonecznienie[78] := -1;
   Naslonecznienie[79] := -1;
   Naslonecznienie[80] := -1;
   Naslonecznienie[81] := -1;
   Naslonecznienie[82] := -1;
   Naslonecznienie[83] := -1;
   Naslonecznienie[84] := -1;
   Naslonecznienie[85] := -1;
   Naslonecznienie[86] := -1;
   Naslonecznienie[87] := -1;
   Naslonecznienie[88] := -1;
   Naslonecznienie[89] := -1;
   Naslonecznienie[90] := -1;
   Naslonecznienie[91] := -1;
   Naslonecznienie[92] := -1;
   Naslonecznienie[93] := -1;
   Naslonecznienie[94] := -1;
   Naslonecznienie[95] := -1;
   Naslonecznienie[96] := -1;
   Naslonecznienie[97] := -1;
   Naslonecznienie[98] := -1;
   Naslonecznienie[99] := -1;
   Naslonecznienie[100] := -1;
   Naslonecznienie[101] := -1;
   Naslonecznienie[102] := -1;
   Naslonecznienie[103] := -1;
   Naslonecznienie[104] := -1;
   Naslonecznienie[105] := -1;
   Naslonecznienie[106] := -1;
   Naslonecznienie[107] := -1;
   Naslonecznienie[108] := -1;
   Naslonecznienie[109] := -1;
   Naslonecznienie[110] := -1;
   Naslonecznienie[111] := -1;
   // Temperatura_srednia[0] : Dzień 1.
END_DATA_BLOCK

// folder: (top level)

ORGANIZATION_BLOCK "Main"   // OB1, LAD, ProgramCycle
TITLE = "Main Program Sweep (Cycle)"
{ S7_Optimized_Access := 'TRUE' }
VERSION : 0.1
   VAR_INPUT
      Initial_Call : Bool;   // Initial call of this OB
      Remanence : Bool;   // =True, if remanent data are available
   END_VAR
BEGIN

REGION Network 1
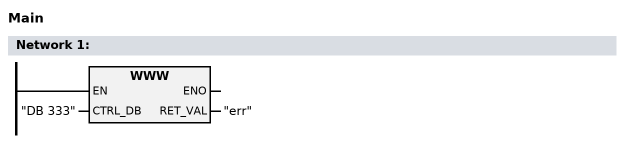
   "err" := WWW(CTRL_DB := "DB 333");
END_REGION
END_ORGANIZATION_BLOCK

(* ===== HMI "HMI_RT_3" =====
system functions are stored by id; their names below are inferred from use
connection "HMI_Connection_4": ETHERNET, SMART_S7_1200_OMS

HMI tags "Default tag table"
   "AlwaysTRUE" : Bool = PLC AlwaysTRUE AT %M1.2, 1 s
   "Grzałka" : Bool = PLC Grzałka AT %Q0.0, 1 s
   "HMI_Aktywacja_trybu_automatycznego" : Bool = PLC HMI.Aktywacja_trybu_automatycznego, 1 s
   "HMI_Aktywacja_trybu_Receptur" : Bool = PLC HMI.Aktywacja_trybu_Receptur, 1 s
   "HMI_Aktywacja_trybu_zapis_Receptur" : Bool = PLC HMI.Aktywacja_trybu_zapis_Receptur, 1 s
   "HMI_Reset_Trybow" : Bool = PLC HMI.Reset_Trybow, 1 s
   "Pompa_podlewanie" : Bool = PLC Pompa_podlewanie AT %Q1.0, 1 s
   "Pompa_zraszacze" : Bool = PLC Pompa_zraszacze AT %Q0.2, 1 s
   "Tag_ScreenNumber" : Int = PLC HMI.Numer_ekranu_HMI AT %MD0, 100 ms
   "Tryb_auto_parametry_Naslonecznienie" : Int = PLC Tryb_auto_parametry.Naslonecznienie, 1 s
   "Tryb_auto_parametry_Stezenie_co2" : Int = PLC Tryb_auto_parametry.Stezenie_co2, 1 s
   "Tryb_auto_parametry_System_okien" : Bool = PLC Tryb_auto_parametry.System_okien, 1 s
   "Tryb_auto_parametry_Temperatura" : Real = PLC Tryb_auto_parametry.Temperatura, 1 s
   "Tryb_auto_parametry_Wilgotnosc_gleby" : Int = PLC Tryb_auto_parametry.Wilgotnosc_gleby, 1 s
   "Tryb_auto_parametry_Wilgotnosc_powietrza" : Int = PLC Tryb_auto_parametry.Wilgotnosc_powietrza, 1 s
   "Wentylator" : Bool = PLC Wentylator AT %Q0.1, 1 s

HMI tags "Z_PLC"
   "Czujnik_wilgotności_powietrza" : Int = PLC Wejscia_PLC.Czujnik_wilgotności_powietrza, 500 ms
   "Temperatura_wewnetrzna" : Real = PLC Wejscia_PLC.Temperatura_wewnetrzna, 500 ms
   "Czujnik_natezenia_światła" : Int = PLC Wejscia_PLC.Czujnik_natezenia_swiatła, 500 ms
   "Czujnik_wilgotności_gleby" : Int = PLC Wejscia_PLC.Czujnik_wilgotności_gleby, 500 ms
   "Wewnetrzny_czujnik_CO2" : Int = PLC Wejscia_PLC.Wewnetrzny_czujnik_CO2, 500 ms
   "Czujnik_wiatru" : Int = PLC Wejscia_PLC.Czujnik_wiatru, 500 ms
   "Stopien_zasloniecia_rolet" : Int = PLC Wejscia_PLC.Stopien_zasloniecia_rolet, 1 s
   "Zewnetrzny_czujnik_CO2" : Int = PLC Wejscia_PLC.Zewnetrzny_czujnik_CO2 AT %DB1.DBW0, 1 s
   "Temperatura_zewnetrzna" : Real = PLC Wejscia_PLC.Temperatura_zewnetrzna AT %DB1.DBW0, 1 s

HMI tags "Do_PLC"
   "System_okien_auto" : Bool = PLC HMI.System_okien_auto, 500 ms
   "Stopien_zasloniecia_rolet_manual" : Int = PLC HMI.Stopien_zasloniecia_rolet_manual, 100 ms
   "Przycisk_zraszania_manual" : Bool = PLC HMI.Przycisk_zraszacze_manual AT %Q0.2, 100 ms
   "Przycisk_wentylacja_manual" : Bool = PLC HMI.Przycisk_wentylacja_manual AT %Q0.1, 100 ms
   "Przycisk_grzanie_manual" : Bool = PLC HMI.Przycisk_grzanie_manual AT %Q0.0, 100 ms
   "Otwarcie_okien_man" : Bool = PLC HMI.Otwarcie_okien_manual AT %DB1.DBW0, 100 ms
   "Temperatura_auto" : Real = PLC HMI.Temperatura_auto, 500 ms
   "Naslonecznienie_auto" : Int = PLC HMI.Naslonecznienie_auto AT %DB1.DBW0, 500 ms
   "Wilgotnosc_powietrza_auto" : Int = PLC HMI.Wilgotnosc_powietrza_auto AT %DB1.DBW0, 500 ms
   "Wilgotnosc_gleby_auto" : Int = PLC HMI.Wilgotnosc_gleby_auto AT %DB1.DBW0, 500 ms
   "Przycisk_zatwierdz_auto" : Bool = PLC HMI.Przycisk_zatwierdz_auto AT %DB1.DBW0, 100 ms
   "nazwa_receptury" : String[254] = PLC HMI.nazwa_receptury AT %DB1.DBX0.0, 500 ms
   "przycisk_zatwierdz_zapis_receptury" : Bool = PLC HMI.Przycisk_zatwierdz_zapis_receptury AT %DB1.DBX0.0, 500 ms
   "HMI_Przycisk_zatwierdz_wybor_receptury" : Bool = PLC HMI.Przycisk_zatwierdz_wybor_receptury AT %DB1.DBX0.0, 500 ms
   "Przycisk_podlewania_manual" : Bool = PLC HMI.Przycisk_podlewanie_manual AT %Q0.2, 100 ms
   "Poziom_CO2_auto" : Int = PLC HMI.Poziom_CO2_auto AT %DB1.DBX0.0, 1 s

analog alarms
   3: 'Podmuchy wiatru osiągają wartości powyżej 35 km/h, system automatyczny zamyka okna.', class Warnings, trigger "Czujnik_wiatru"
   2: 'Temperatura powyżej 35 stopni / Temperatura powyżej 35 stopni, zaleca się wyłączenie grzania.', class Warnings, trigger "Temperatura_wewnetrzna"
   5: 'Temperatura powyżej 45 stopni, NIEZWŁOCZNIE SPRAWDŹ DZIAŁANIE GRZAŁKI, TERMOMETRU LUB WENTYLATORA. / Temperatura powyżej 45 stopni, NIEZWŁOCZNIE SPRAWDŹ DZIAŁANIE GRZAŁKI, TERMOMETRU LUB WENTYLATORA. JEŚLI TEMPERATURA NIE SPADA ZALECA SIĘ EWAKUOWAĆ WSZYSTKICH PRZEBYWAJĄCYCH W POMIESZCZENIU', class Errors, trigger "Temperatura_wewnetrzna"
   4: 'Stężenie CO2 ma powyżej 5000 jednostek. NIEZWŁOCZNIE OTWORZ OKNA ORAZ ZAŁĄCZ WENTYLATOR, NASTĘPNIE NALEŻY EWAKUOWAĆ WSZYSTKUCH ZNAJDUJĄCYCH SIĘ W POMIESZCZENIU / Stężenie CO2 ma powyżej 5000 jednostek. NIEZWŁOCZNIE OTWORZ OKNA ORAZ ZAŁĄCZ WENTYLATOR, NASTĘPNIE NALEŻY EWAKUOWAĆ WSZYSTKUCH ZNAJDUJĄCYCH SIĘ W POMIESZCZENIU', class Errors, trigger "Wewnetrzny_czujnik_CO2"
   1: 'Stężenie CO2 ma powyżej 3000 jednostek / Stężenie CO2 ma powyżej 3000 jednostek, dłużesze przebywanie w takim środowisku może być szkodliwe dla człowieka. Zalecane jest włączenie wentylacji lub otworzenie okien.', class Warnings, trigger "Wewnetrzny_czujnik_CO2"

text list "receptury": 0..1 ''

recipe "Receptura_nr1": Temperatura <- "Tryb_auto_parametry_Temperatura", Wilgotność Powietrza <- "Tryb_auto_parametry_Wilgotnosc_powietrza", Wilgotność gleby <- "Tryb_auto_parametry_Wilgotnosc_gleby", System okien <- "Tryb_auto_parametry_System_okien", Stężenie CO2 <- "Tryb_auto_parametry_Stezenie_co2", Nasłonecznienie <- "Tryb_auto_parametry_Naslonecznienie"

